REGION Network 2
   RUNG wire#powerrail
      { S7_Templates := "SrcType := Byte" } EQ_Contact(in1 := #Lbyte, in2 := 16#00)
      wire#w1
      Coil( #工作正常 )
   END_RUNG
   RUNG wire#w1
      Coil( #Error.%X1 )
   END_RUNG
   // the same network as SCL:
   #工作正常 := #Lbyte = 16#00;
   #Error.%X1 := #工作正常;
END_REGION

REGION Network 3
   RUNG wire#powerrail
      { S7_Templates := "SrcType := Byte" } EQ_Contact(in1 := #Lbyte, in2 := 16#01)
      wire#w1
      Coil( #无反馈信号 )
   END_RUNG
   RUNG wire#w1
      Coil( #Error.%X2 )
   END_RUNG
   // the same network as SCL:
   #无反馈信号 := #Lbyte = 16#01;
   #Error.%X2 := #无反馈信号;
END_REGION

REGION Network 4
   RUNG wire#powerrail
      { S7_Templates := "SrcType := Byte" } EQ_Contact(in1 := #Lbyte, in2 := 16#02)
      wire#w1
      Coil( #欠压保护 )
   END_RUNG
   RUNG wire#w1
      Coil( #Error.%X3 )
   END_RUNG
   // the same network as SCL:
   #欠压保护 := #Lbyte = 16#02;
   #Error.%X3 := #欠压保护;
END_REGION

REGION Network 5
   RUNG wire#powerrail
      { S7_Templates := "SrcType := Byte" } EQ_Contact(in1 := #Lbyte, in2 := 16#03)
      wire#w1
      Coil( #过压保护 )
   END_RUNG
   RUNG wire#w1
      Coil( #Error.%X4 )
   END_RUNG
   // the same network as SCL:
   #过压保护 := #Lbyte = 16#03;
   #Error.%X4 := #过压保护;
END_REGION

REGION Network 6
   RUNG wire#powerrail
      { S7_Templates := "SrcType := Byte" } EQ_Contact(in1 := #Lbyte, in2 := 16#04)
      wire#w1
      Coil( #过流保护 )
   END_RUNG
   RUNG wire#w1
      Coil( #Error.%X5 )
   END_RUNG
   // the same network as SCL:
   #过流保护 := #Lbyte = 16#04;
   #Error.%X5 := #过流保护;
END_REGION

REGION Network 7
   RUNG wire#powerrail
      { S7_Templates := "SrcType := Byte" } EQ_Contact(in1 := #Lbyte, in2 := 16#05)
      wire#w1
      Coil( #过温保护 )
   END_RUNG
   RUNG wire#w1
      Coil( #Error.%X6 )
   END_RUNG
   // the same network as SCL:
   #过温保护 := #Lbyte = 16#05;
   #Error.%X6 := #过温保护;
END_REGION

REGION Network 8
   RUNG wire#powerrail
      { S7_Templates := "SrcType := Byte" } EQ_Contact(in1 := #Lbyte, in2 := 16#06)
      wire#w1
      Coil( #磁控管故障 )
   END_RUNG
   RUNG wire#w1
      Coil( #Error.%X7 )
   END_RUNG
   // the same network as SCL:
   #磁控管故障 := #Lbyte = 16#06;
   #Error.%X7 := #磁控管故障;
END_REGION

REGION Network 9
   RUNG wire#powerrail
      { S7_Templates := "SrcType := Byte" } EQ_Contact(in1 := #Lbyte, in2 := 16#07)
      wire#w1
      Coil( #浪涌保护 )
   END_RUNG
   RUNG wire#w1
      Coil( #Error.%X8 )
   END_RUNG
   // the same network as SCL:
   #浪涌保护 := #Lbyte = 16#07;
   #Error.%X8 := #浪涌保护;
END_REGION

REGION Network 10
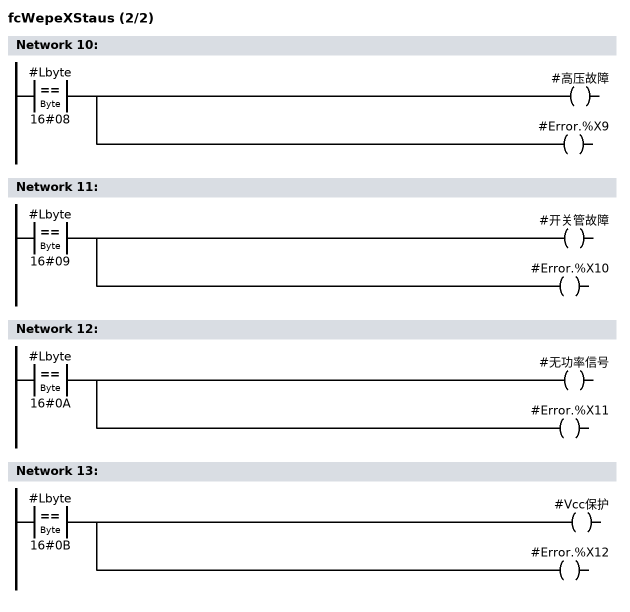
   RUNG wire#powerrail
      { S7_Templates := "SrcType := Byte" } EQ_Contact(in1 := #Lbyte, in2 := 16#08)
      wire#w1
      Coil( #高压故障 )
   END_RUNG
   RUNG wire#w1
      Coil( #Error.%X9 )
   END_RUNG
   // the same network as SCL:
   #高压故障 := #Lbyte = 16#08;
   #Error.%X9 := #高压故障;
END_REGION

REGION Network 11
   RUNG wire#powerrail
      { S7_Templates := "SrcType := Byte" } EQ_Contact(in1 := #Lbyte, in2 := 16#09)
      wire#w1
      Coil( #开关管故障 )
   END_RUNG
   RUNG wire#w1
      Coil( #Error.%X10 )
   END_RUNG
   // the same network as SCL:
   #开关管故障 := #Lbyte = 16#09;
   #Error.%X10 := #开关管故障;
END_REGION

REGION Network 12
   RUNG wire#powerrail
      { S7_Templates := "SrcType := Byte" } EQ_Contact(in1 := #Lbyte, in2 := 16#0A)
      wire#w1
      Coil( #无功率信号 )
   END_RUNG
   RUNG wire#w1
      Coil( #Error.%X11 )
   END_RUNG
   // the same network as SCL:
   #无功率信号 := #Lbyte = 16#0A;
   #Error.%X11 := #无功率信号;
END_REGION

REGION Network 13
   RUNG wire#powerrail
      { S7_Templates := "SrcType := Byte" } EQ_Contact(in1 := #Lbyte, in2 := 16#0B)
      wire#w1
      Coil( #Vcc保护 )
   END_RUNG
   RUNG wire#w1
      Coil( #Error.%X12 )
   END_RUNG
   // the same network as SCL:
   #Vcc保护 := #Lbyte = 16#0B;
   #Error.%X12 := #Vcc保护;
END_REGION
END_FUNCTION

FUNCTION "fcInt_to_mTime" : Void   // FC103, LAD
{ S7_Optimized_Access := 'TRUE' }
VERSION : 0.1
   VAR_INPUT
      intData : Int;
   END_VAR
   VAR_OUTPUT
      mTimeData : Time;
      sTimeData : Time;
   END_VAR
   VAR_TEMP
      dintData1 : DInt;
      dintData2 : DInt;
      dintData3 : DInt;
   END_VAR
BEGIN

REGION Network 1
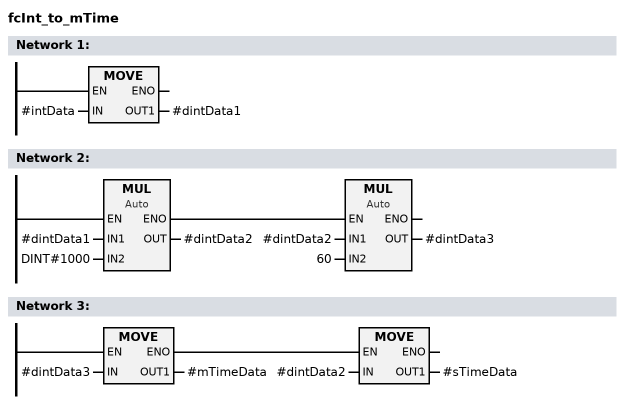
   RUNG wire#powerrail
      Move(in := #intData, out1 => #dintData1)
   END_RUNG
   // the same network as SCL:
   #dintData1 := #intData;
END_REGION

REGION Network 2
   RUNG wire#powerrail
      Mul(in1 := #dintData1, in2 := DINT#1000, out => #dintData2)
      Mul(in1 := #dintData2, in2 := 60, out => #dintData3)
   END_RUNG
   // the same network as SCL:
   #dintData2 := #dintData1 * DINT#1000;
   #dintData3 := #dintData2 * 60;
END_REGION

REGION Network 3
   RUNG wire#powerrail
      Move(in := #dintData3, out1 => #mTimeData)
      Move(in := #dintData2, out1 => #sTimeData)
   END_RUNG
   // the same network as SCL:
   #mTimeData := #dintData3;
   #sTimeData := #dintData2;
END_REGION
END_FUNCTION

FUNCTION "fcArray_Int_mTime" : Void   // FC104, LAD
{ S7_Optimized_Access := 'TRUE' }
VERSION : 0.1
   VAR_INPUT
      "Int" : Array[1..16] of Int;
   END_VAR
   VAR_OUTPUT
      mTimeOut : Array[1..16] of Time;
      sTimeOut : Array[1..16] of Time;
   END_VAR
   VAR_TEMP   // added for the SCL form of the ladder/FBD networks
      _w1 : Bool;
      _w2 : Bool;
      _w3 : Bool;
   END_VAR
BEGIN

REGION Network 1
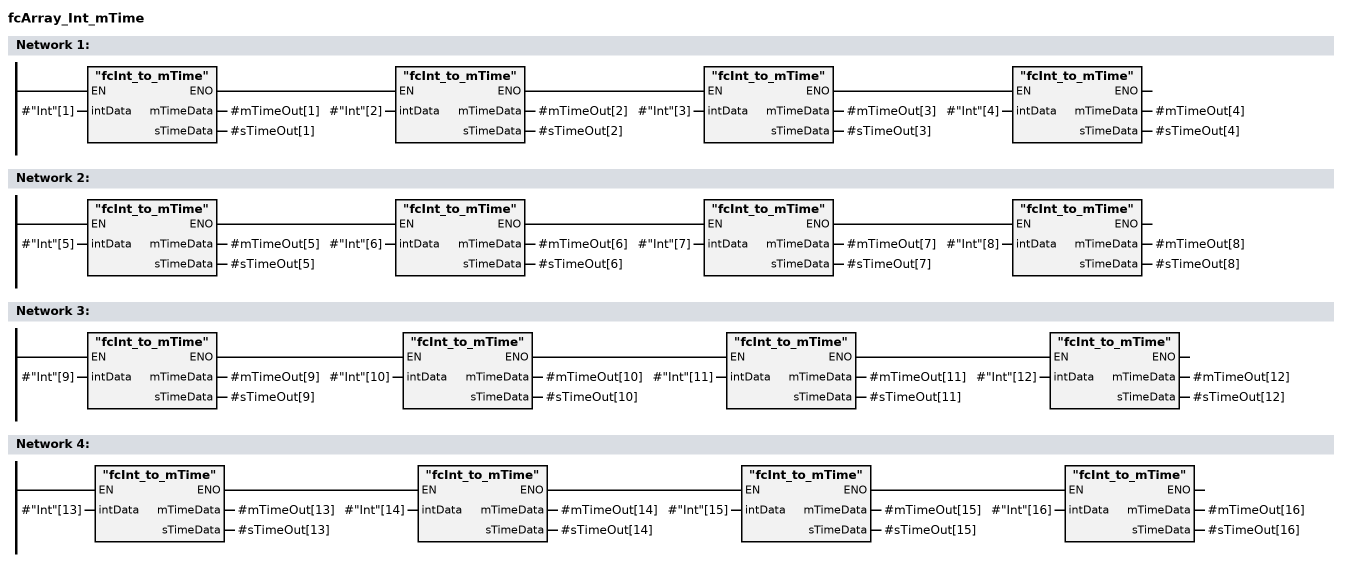
   RUNG wire#powerrail
      "fcInt_to_mTime"(intData := #"Int"[1], mTimeData => #mTimeOut[1], sTimeData => #sTimeOut[1])
      "fcInt_to_mTime"(intData := #"Int"[2], mTimeData => #mTimeOut[2], sTimeData => #sTimeOut[2])
      "fcInt_to_mTime"(intData := #"Int"[3], mTimeData => #mTimeOut[3], sTimeData => #sTimeOut[3])
      "fcInt_to_mTime"(intData := #"Int"[4], mTimeData => #mTimeOut[4], sTimeData => #sTimeOut[4])
   END_RUNG
   // the same network as SCL:
   "fcInt_to_mTime"(intData := #"Int"[1], mTimeData => #mTimeOut[1], sTimeData => #sTimeOut[1], ENO => #_w1);
   "fcInt_to_mTime"(EN := #_w1,
                    intData := #"Int"[2],
                    mTimeData => #mTimeOut[2],
                    sTimeData => #sTimeOut[2],
                    ENO => #_w2);
   "fcInt_to_mTime"(EN := #_w2,
                    intData := #"Int"[3],
                    mTimeData => #mTimeOut[3],
                    sTimeData => #sTimeOut[3],
                    ENO => #_w3);
   IF #_w3 THEN
       "fcInt_to_mTime"(intData := #"Int"[4], mTimeData => #mTimeOut[4], sTimeData => #sTimeOut[4]);
   END_IF;
END_REGION

REGION Network 2
   RUNG wire#powerrail
      "fcInt_to_mTime"(intData := #"Int"[5], mTimeData => #mTimeOut[5], sTimeData => #sTimeOut[5])
      "fcInt_to_mTime"(intData := #"Int"[6], mTimeData => #mTimeOut[6], sTimeData => #sTimeOut[6])
      "fcInt_to_mTime"(intData := #"Int"[7], mTimeData => #mTimeOut[7], sTimeData => #sTimeOut[7])
      "fcInt_to_mTime"(intData := #"Int"[8], mTimeData => #mTimeOut[8], sTimeData => #sTimeOut[8])
   END_RUNG
   // the same network as SCL:
   "fcInt_to_mTime"(intData := #"Int"[5], mTimeData => #mTimeOut[5], sTimeData => #sTimeOut[5], ENO => #_w1);
   "fcInt_to_mTime"(EN := #_w1,
                    intData := #"Int"[6],
                    mTimeData => #mTimeOut[6],
                    sTimeData => #sTimeOut[6],
                    ENO => #_w2);
   "fcInt_to_mTime"(EN := #_w2,
                    intData := #"Int"[7],
                    mTimeData => #mTimeOut[7],
                    sTimeData => #sTimeOut[7],
                    ENO => #_w3);
   IF #_w3 THEN
       "fcInt_to_mTime"(intData := #"Int"[8], mTimeData => #mTimeOut[8], sTimeData => #sTimeOut[8]);
   END_IF;
END_REGION

REGION Network 3
   RUNG wire#powerrail
      "fcInt_to_mTime"(intData := #"Int"[9], mTimeData => #mTimeOut[9], sTimeData => #sTimeOut[9])
      "fcInt_to_mTime"(intData := #"Int"[10], mTimeData => #mTimeOut[10], sTimeData => #sTimeOut[10])
      "fcInt_to_mTime"(intData := #"Int"[11], mTimeData => #mTimeOut[11], sTimeData => #sTimeOut[11])
      "fcInt_to_mTime"(intData := #"Int"[12], mTimeData => #mTimeOut[12], sTimeData => #sTimeOut[12])
   END_RUNG
   // the same network as SCL:
   "fcInt_to_mTime"(intData := #"Int"[9], mTimeData => #mTimeOut[9], sTimeData => #sTimeOut[9], ENO => #_w1);
   "fcInt_to_mTime"(EN := #_w1,
                    intData := #"Int"[10],
                    mTimeData => #mTimeOut[10],
                    sTimeData => #sTimeOut[10],
                    ENO => #_w2);
   "fcInt_to_mTime"(EN := #_w2,
                    intData := #"Int"[11],
                    mTimeData => #mTimeOut[11],
                    sTimeData => #sTimeOut[11],
                    ENO => #_w3);
   IF #_w3 THEN
       "fcInt_to_mTime"(intData := #"Int"[12], mTimeData => #mTimeOut[12], sTimeData => #sTimeOut[12]);
   END_IF;
END_REGION

REGION Network 4
   RUNG wire#powerrail
      "fcInt_to_mTime"(intData := #"Int"[13], mTimeData => #mTimeOut[13], sTimeData => #sTimeOut[13])
      "fcInt_to_mTime"(intData := #"Int"[14], mTimeData => #mTimeOut[14], sTimeData => #sTimeOut[14])
      "fcInt_to_mTime"(intData := #"Int"[15], mTimeData => #mTimeOut[15], sTimeData => #sTimeOut[15])
      "fcInt_to_mTime"(intData := #"Int"[16], mTimeData => #mTimeOut[16], sTimeData => #sTimeOut[16])
   END_RUNG
   // the same network as SCL:
   "fcInt_to_mTime"(intData := #"Int"[13], mTimeData => #mTimeOut[13], sTimeData => #sTimeOut[13], ENO => #_w1);
   "fcInt_to_mTime"(EN := #_w1,
                    intData := #"Int"[14],
                    mTimeData => #mTimeOut[14],
                    sTimeData => #sTimeOut[14],
                    ENO => #_w2);
   "fcInt_to_mTime"(EN := #_w2,
                    intData := #"Int"[15],
                    mTimeData => #mTimeOut[15],
                    sTimeData => #sTimeOut[15],
                    ENO => #_w3);
   IF #_w3 THEN
       "fcInt_to_mTime"(intData := #"Int"[16], mTimeData => #mTimeOut[16], sTimeData => #sTimeOut[16]);
   END_IF;
END_REGION
END_FUNCTION

FUNCTION "fcArray_bool_to_bool" : Void   // FC105, LAD
{ S7_Optimized_Access := 'TRUE' }
VERSION : 0.1
   VAR_INPUT
      In : Array[1..16] of Bool;
   END_VAR
   VAR_OUTPUT
      Out : Bool;
   END_VAR
BEGIN

REGION Network 1
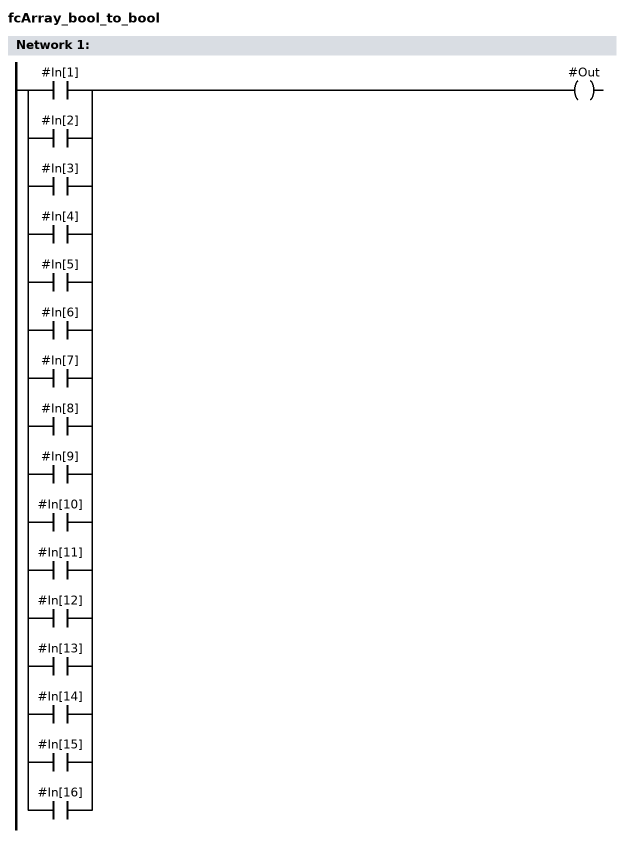
   RUNG wire#powerrail
      Contact( #In[1] )
      wire#w1
      Coil( #Out )
   END_RUNG
   RUNG wire#powerrail
      Contact( #In[2] )
   END_RUNG wire#w1
   RUNG wire#powerrail
      Contact( #In[3] )
   END_RUNG wire#w1
   RUNG wire#powerrail
      Contact( #In[4] )
   END_RUNG wire#w1
   RUNG wire#powerrail
      Contact( #In[5] )
   END_RUNG wire#w1
   RUNG wire#powerrail
      Contact( #In[6] )
   END_RUNG wire#w1
   RUNG wire#powerrail
      Contact( #In[7] )
   END_RUNG wire#w1
   RUNG wire#powerrail
      Contact( #In[8] )
   END_RUNG wire#w1
   RUNG wire#powerrail
      Contact( #In[9] )
   END_RUNG wire#w1
   RUNG wire#powerrail
      Contact( #In[10] )
   END_RUNG wire#w1
   RUNG wire#powerrail
      Contact( #In[11] )
   END_RUNG wire#w1
   RUNG wire#powerrail
      Contact( #In[12] )
   END_RUNG wire#w1
   RUNG wire#powerrail
      Contact( #In[13] )
   END_RUNG wire#w1
   RUNG wire#powerrail
      Contact( #In[14] )
   END_RUNG wire#w1
   RUNG wire#powerrail
      Contact( #In[15] )
   END_RUNG wire#w1
   RUNG wire#powerrail
      Contact( #In[16] )
   END_RUNG wire#w1
   // the same network as SCL:
   #Out := #In[1] OR #In[2] OR #In[3] OR #In[4] OR #In[5] OR #In[6] OR #In[7] OR #In[8] OR #In[9] OR #In[10] OR #In[11] OR #In[12] OR #In[13] OR #In[14] OR #In[15] OR #In[16];
END_REGION
END_FUNCTION

ORGANIZATION_BLOCK "Main"   // OB1, LAD, ProgramCycle
TITLE = "Main Program Sweep (Cycle)"
{ S7_Optimized_Access := 'TRUE' }
VERSION : 0.1
   VAR_INPUT
      Initial_Call : Bool;   // Initial call of this OB
      Remanence : Bool;   // =True, if remanent data are available
   END_VAR
BEGIN

REGION Network 1
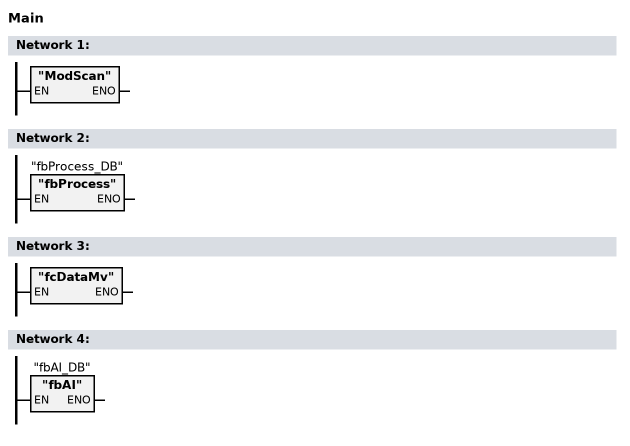
   RUNG wire#powerrail
      "ModScan"()
   END_RUNG
   // the same network as SCL:
   "ModScan"();
END_REGION

REGION Network 2
   RUNG wire#powerrail
      "fbProcess_DB"()
   END_RUNG
   // the same network as SCL:
   "fbProcess_DB"();   // "fbProcess"
END_REGION

REGION Network 3
   RUNG wire#powerrail
      "fcDataMv"()
   END_RUNG
   // the same network as SCL:
   "fcDataMv"();
END_REGION

REGION Network 4
   RUNG wire#powerrail
      "fbAI_DB"()
   END_RUNG
   // the same network as SCL:
   "fbAI_DB"();   // "fbAI"
END_REGION
END_ORGANIZATION_BLOCK

// folder: System blocks/Program resources

FUNCTION "ModScan" : Void   // FC10000, LAD
TITLE = ModScan
{ S7_Optimized_Access := 'TRUE' }
AUTHOR : SIMATIC
VERSION : 4.0
BEGIN

REGION Network 1: Modbus-RTU Job scan
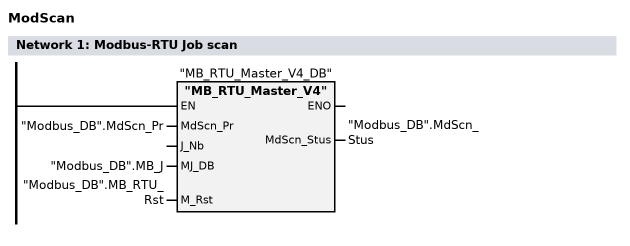
   RUNG wire#powerrail
      "MB_RTU_Master_V4_DB"(MdScn_Pr := "Modbus_DB".MdScn_Pr, J_Nb :=, MJ_DB := "Modbus_DB".MB_J, M_Rst := "Modbus_DB".MB_RTU_Rst, MdScn_Stus => "Modbus_DB".MdScn_Stus)
   END_RUNG
   // the same network as SCL:
   "MB_RTU_Master_V4_DB"(MdScn_Pr := "Modbus_DB".MdScn_Pr,   // "MB_RTU_Master_V4"
                         MJ_DB := "Modbus_DB".MB_J,
                         M_Rst := "Modbus_DB".MB_RTU_Rst,
                         MdScn_Stus => "Modbus_DB".MdScn_Stus);
END_REGION
END_FUNCTION

(* ===== HMI "HMI_RT_1" =====
system functions are stored by id; their names below are inferred from use
connection "HMI_连接_1": ETHERNET, SMART_S7_1200_OMS

HMI tags "变量表_1"
   "WepeX_PowerSPCom" : Int = PLC dbHMI.WepeX_PowerSPCom AT %DB50.DBW0, 1 s
   "WepeX_ActpowerCom" : Int = PLC dbHMI.WepeX_ActpowerCom AT %DB50.DBW38, 1 s
   "Mode" : Bool = PLC dbHMI.Mode AT %DB50.DBX164.0, 1 s
   "WepeX_PowerMan" : Bool = PLC dbHMI.WepeX_PowerMan AT %DB50.DBX164.1, 1 s
   "CoolingWaterMan" : Bool = PLC dbHMI.CoolingWaterMan AT %DB50.DBX164.2, 1 s
   "AirCompressorMan" : Bool = PLC dbHMI.AirCompressorMan AT %DB50.DBX164.3, 1 s
   "BlowerMan" : Bool = PLC dbHMI.BlowerMan AT %DB50.DBX164.4, 1 s
   "PeristalticpumpMan" : Bool = PLC dbHMI.PeristalticpumpMan AT %DB50.DBX164.5, 1 s
   "1YV1Man" : Bool = PLC dbHMI.1YV1Man AT %DB50.DBX164.6, 1 s
   "1YV2Man" : Bool = PLC dbHMI.1YV2Man AT %DB50.DBX164.7, 1 s
   "2YV1Man" : Bool = PLC dbHMI.2YV1Man AT %DB50.DBX165.0, 1 s
   "2YV2Man" : Bool = PLC dbHMI.2YV2Man AT %DB50.DBX165.1, 1 s
   "WepeXP1通信正常" : Bool = PLC dbHMI.WepeXP1通信正常 AT %DB50.DBX170.0, 1 s
   "WepeXP1通信不正常" : Bool = PLC dbHMI.WepeXP1通信不正常 AT %DB50.DBX170.1, 1 s
   "WepeXP1工作正常" : Bool = PLC dbHMI.WepeXP1工作正常 AT %DB50.DBX170.2, 1 s
   "WepeXP1无反馈信号" : Bool = PLC dbHMI.WepeXP1无反馈信号 AT %DB50.DBX170.3, 1 s
   "WepeXP1欠压保护" : Bool = PLC dbHMI.WepeXP1欠压保护 AT %DB50.DBX170.4, 1 s
   "WepeXP1过压保护" : Bool = PLC dbHMI.WepeXP1过压保护 AT %DB50.DBX170.5, 1 s
   "WepeXP1过流保护" : Bool = PLC dbHMI.WepeXP1过流保护 AT %DB50.DBX170.6, 1 s
   "WepeXP1过温保护" : Bool = PLC dbHMI.WepeXP1过温保护 AT %DB50.DBX170.7, 1 s
   "WepeXP1磁控管故障" : Bool = PLC dbHMI.WepeXP1磁控管故障 AT %DB50.DBX171.0, 1 s
   "WepeXP1浪涌保护" : Bool = PLC dbHMI.WepeXP1浪涌保护 AT %DB50.DBX171.1, 1 s
   "WepeXP1高压故障" : Bool = PLC dbHMI.WepeXP1高压故障 AT %DB50.DBX171.2, 1 s
   "WepeXP1开关管故障" : Bool = PLC dbHMI.WepeXP1开关管故障 AT %DB50.DBX171.3, 1 s
   "WepeXP1无功率信号" : Bool = PLC dbHMI.WepeXP1无功率信号 AT %DB50.DBX171.4, 1 s
   "WepeXP1Vcc保护" : Bool = PLC dbHMI.WepeXP1Vcc保护 AT %DB50.DBX171.5, 1 s
   "WepeXP1通信状态" : Int = PLC dbHMI.WepeXP1通信状态 AT %DB50.DBW172, 1 s
   "微波状态" : Int = PLC dbHMI.微波状态 AT %DB50.DBW174, 1 s
   "火炬状态" : Int = PLC dbHMI.火炬状态 AT %DB50.DBW176, 1 s
   "Start" : Bool = PLC dbHMI.Start AT %DB50.DBX178.0, 1 s
   "Stop" : Bool = PLC dbHMI.Stop AT %DB50.DBX178.1, 1 s
   "Reset" : Bool = PLC dbHMI.Reset AT %DB50.DBX178.2, 1 s
   "Running" : Bool = PLC dbHMI.Running AT %DB50.DBX178.3, 1 s
   "WepeXPowerOut" : Bool = PLC WepeXEnable AT %Q0.1, 1 s
   "CoolingWater" : Bool = PLC CoolingWater AT %Q0.2, 1 s
   "Blower" : Bool = PLC Blower AT %Q0.3, 1 s
   "AirCompressor" : Bool = PLC AirCompressor AT %Q0.4, 1 s
   "Peristalticpump" : Bool = PLC Peristalticpump AT %Q0.0, 1 s
   "气体温度" : Real = PLC dbHMI.气体温度 AT %DB50.DBD180, 1 s
   "1YV1" : Bool = PLC 1YV1 AT %Q1.0, 1 s
   "1YV2" : Bool = PLC 1YV2 AT %Q1.1, 1 s
   "2YV1" : Bool = PLC 2YV1 AT %Q1.2, 1 s
   "2YV2" : Bool = PLC 2YV2 AT %Q1.3, 1 s
   "3YV1Man" : Bool = PLC dbHMI.3YV1Man AT %DB50.DBX165.2, 1 s
   "3YV1" : Bool = PLC 3YV1 AT %Q1.4, 1 s
   "3YV2Man" : Bool = PLC dbHMI.3YV2Man AT %DB50.DBX165.3, 1 s
   "3YV2" : Bool = PLC 3YV2 AT %Q1.5, 1 s
   "4YVMan" : Bool = PLC dbHMI.4YVMan AT %DB50.DBX165.4, 1 s
   "4YV" : Bool = PLC 4YV AT %Q1.6, 1 s
   "inUnit.Coolingwater" : Bool = PLC dbHMI.inUnit.Coolingwater AT %DB50.DBX184.0, 1 s
   "inUnit.AirCompressor" : Bool = PLC dbHMI.inUnit.AirCompressor AT %DB50.DBX184.1, 1 s
   "inUnit.Peristalticpump" : Bool = PLC dbHMI.inUnit.Peristalticpump AT %DB50.DBX184.2, 1 s
   "inUnit.WepeX_Enable" : Bool = PLC dbHMI.inUnit.WepeX_Enable AT %DB50.DBX184.3, 1 s
   "inUnit.AYV1" : Bool = PLC dbHMI.inUnit.AYV1 AT %DB50.DBX184.4, 1 s
   "inUnit.AYV2" : Bool = PLC dbHMI.inUnit.AYV2 AT %DB50.DBX184.5, 1 s
   "inUnit.BYV1" : Bool = PLC dbHMI.inUnit.BYV1 AT %DB50.DBX184.6, 1 s
   "inUnit.BYV2" : Bool = PLC dbHMI.inUnit.BYV2 AT %DB50.DBX184.7, 1 s
   "inUnit.CYV1" : Bool = PLC dbHMI.inUnit.CYV1 AT %DB50.DBX185.0, 1 s
   "inUnit.CYV2" : Bool = PLC dbHMI.inUnit.CYV2 AT %DB50.DBX185.1, 1 s
   "inUnit.DYV" : Bool = PLC dbHMI.inUnit.DYV AT %DB50.DBX185.2, 1 s
   "inUnit.Blower" : Bool = PLC dbHMI.inUnit.Blower AT %DB50.DBX185.3, 1 s
   "inUnit.Runtime" : Int = PLC dbHMI.inUnit.Runtime AT %DB50.DBW186, 1 s
   "inUnit.WepeX_Power" : Int = PLC dbHMI.inUnit.WepeX_Power AT %DB50.DBW188, 1 s
   "inUnit.Donebit" : Int = PLC dbHMI.inUnit.Donebit AT %DB50.DBW190, 1 s
   "ActUnit.Coolingwater" : Bool = PLC dbHMI.ActRcpUnit.Coolingwater AT %DB50.DBX202.0, 1 s
   "ActUnit.AirCompressor" : Bool = PLC dbHMI.ActRcpUnit.AirCompressor AT %DB50.DBX202.1, 1 s
   "ActUnit.Peristalticpump" : Bool = PLC dbHMI.ActRcpUnit.Peristalticpump AT %DB50.DBX202.2, 1 s
   "ActUnit.WepeX_Enable" : Bool = PLC dbHMI.ActRcpUnit.WepeX_Enable AT %DB50.DBX202.3, 1 s
   "ActUnit.AYV1" : Bool = PLC dbHMI.ActRcpUnit.AYV1 AT %DB50.DBX202.4, 1 s
   "ActUnit.AYV2" : Bool = PLC dbHMI.ActRcpUnit.AYV2 AT %DB50.DBX202.5, 1 s
   "ActUnit.BYV1" : Bool = PLC dbHMI.ActRcpUnit.BYV1 AT %DB50.DBX202.6, 1 s
   "ActUnit.BYV2" : Bool = PLC dbHMI.ActRcpUnit.BYV2 AT %DB50.DBX202.7, 1 s
   "ActUnit.CYV1" : Bool = PLC dbHMI.ActRcpUnit.CYV1 AT %DB50.DBX203.0, 1 s
   "ActUnit.CYV2" : Bool = PLC dbHMI.ActRcpUnit.CYV2 AT %DB50.DBX203.1, 1 s
   "ActUnit.DYV" : Bool = PLC dbHMI.ActRcpUnit.DYV AT %DB50.DBX203.2, 1 s
   "ActUnit.Blower" : Bool = PLC dbHMI.ActRcpUnit.Blower AT %DB50.DBX203.3, 1 s
   "ActUnit.Runtime" : Int = PLC dbHMI.ActRcpUnit.Runtime AT %DB50.DBW204, 1 s
   "ActUnit.WepeX_Power" : Int = PLC dbHMI.ActRcpUnit.WepeX_Power AT %DB50.DBW206, 1 s
   "ActUnit.Donebit" : Int = PLC dbHMI.ActRcpUnit.Donebit AT %DB50.DBW208, 1 s
   "RecipeNum" : Int = PLC dbHMI.RecipeNum AT %DB50.DBW192, 1 s
   "StepNumMan" : Int = PLC dbHMI.StepNumMan AT %DB50.DBW194, 1 s
   "Editor" : Bool = PLC dbHMI.Editor AT %DB50.DBX200.0, 1 s
   "Save" : Bool = PLC dbHMI.Save AT %DB50.DBX200.1, 1 s

discrete alarms
   1: '', class Errors

Template "模板_1" 800x480
   Button "模板_按钮_1" at 0,448 size 96x32; TextOff '自动页面'
      on Click: ActivateScreen("1自动画面", 0)
   Button "模板_按钮_2" at 96,448 size 96x32; TextOff '手动页面'
      on Click: ActivateScreen("2手动画面", 0)
   Button "模板_按钮_3" at 192,448 size 96x32; TextOff '程序设置'
      on Click: ActivateScreen("3程序设置", 0)
   Button "模板_按钮_4" at 288,448 size 96x32; TextOff '温度曲线'
      on Click: ActivateScreen("4温度曲线", 0)
   Button "模板_按钮_5" at 384,448 size 96x32; TextOff '报警信息'
      Appearance <- "Mode"
      on Click: ActivateScreen("5报警信息", 0)
   Button "模板_按钮_6" at 480,448 size 96x32; TextOff '自/手模式'
      on Press: InvertBit("Mode")
      Appearance <- "Mode"

screen "1自动画面" 800x480, template "模板_1"
   TextField "文本域_16" at 73,86 size 57x16; Text '设备状态'
   TextField "文本域_17" at 103,145 size 31x16; Text '微波'
   TextField "文本域_18" at 103,177 size 31x16; Text '火炬'
   TextField "文本域_19" at 103,113 size 31x16; Text '通信'
   TextField "文本域_20" at 102,211 size 31x16; Text '过流'
   TextField "文本域_21" at 102,245 size 31x16; Text '欠流'
   TextField "文本域_22" at 102,280 size 31x16; Text '超温'
   TextField "文本域_14" at 325,75 size 73x20; Text '程序选择'
   Button "按钮_1" at 316,114 size 97x32; TextOff '开放式'
   Button "按钮_2" at 316,187 size 97x32; TextOff '管道式'
   Button "按钮_3" at 314,259 size 97x32; TextOff '自定义'
   Button "按钮_7" at 153,343 size 81x70; TextOff '启动'
      on Press: SetBit("Start")
      on Release: ResetBit("Start")
      Appearance <- "Running"
   TextField "文本域_6" at 575,199 size 73x20; Text '气体余量'
   IOField "I/O 域_4" at 646,191 size 96x32; FormatPattern 9999999
   TextField "文本域_7" at 576,95 size 73x20; Text '实际功率'
   IOField "I/O 域_5" at 648,90 size 96x32; FormatPattern s99999
      ProcessValue <- "WepeX_ActpowerCom"
   TextField "文本域_8" at 745,94 size 16x23; Text 'W'
   TextField "文本域_9" at 575,149 size 73x20; Text '气体温度'
   IOField "I/O 域_6" at 648,141 size 96x32; FormatPattern s999.99
      ProcessValue <- "气体温度"
   TextField "文本域_10" at 745,147 size 25x23; Text '℃'
   Button "按钮_8" at 382,348 size 80x68; TextOff '停止'
      on Press: SetBit("Stop")
      on Release: ResetBit("Stop")
   TextField "文本域_1" at 237,14 size 275x33; Text '多功能等离子消毒机'
   Circle "圆_1" at 74,112 size 20x20
      Appearance <- "WepeXP1通信不正常"
   Circle "圆_2" at 74,144 size 20x20
      Appearance <- "微波状态"
   Circle "圆_3" at 74,177 size 20x20
      Appearance <- "火炬状态"
   Circle "圆_4" at 74,210 size 20x20
      Appearance <- "WepeXP1过流保护"
   Circle "圆_5" at 74,243 size 20x20
      Appearance <- "WepeXP1欠压保护"
   Circle "圆_6" at 74,277 size 20x20
      Appearance <- "WepeXP1过温保护"
   Button "按钮_9" at 606,349 size 82x64; TextOff '复位'
      on Press: SetBit("Reset")
      on Release: ResetBit("Reset")
   TextField "文本域_4" at 749,197 size 16x23; Text '%'

screen "2手动画面" 800x480, template "模板_1"
   Button "按钮_1" at 169,84 size 80x55; TextOff '冷水机'
      on Press: InvertBit("CoolingWaterMan")
      Appearance <- "CoolingWaterMan"
   Button "按钮_2" at 169,258 size 80x55; TextOff '空压机'
      on Press: InvertBit("AirCompressorMan")
      Appearance <- "AirCompressorMan"
   Button "按钮_3" at 169,170 size 80x55; TextOff '风机'
      on Press: InvertBit("BlowerMan")
      Appearance <- "BlowerMan"
   Button "按钮_4" at 169,348 size 80x55; TextOff '蠕动泵'
      on Press: InvertBit("PeristalticpumpMan")
      Appearance <- "PeristalticpumpMan"
   TextField "文本域_6" at 617,102 size 73x20; Text '功率设置'
   IOField "I/O 域_4" at 697,95 size 64x32; FormatPattern 9999
      ProcessValue <- "WepeX_PowerSPCom"
   TextField "文本域_7" at 620,156 size 73x20; Text '实际功率'
   IOField "I/O 域_5" at 700,149 size 57x32; FormatPattern 9999
      ProcessValue <- "WepeX_ActpowerCom"
   TextField "文本域_8" at 764,154 size 16x23; Text 'W'
   TextField "文本域_9" at 620,210 size 73x20; Text '气体余量'
   IOField "I/O 域_6" at 695,205 size 63x32; FormatPattern 999
   TextField "文本域_10" at 755,269 size 25x23; Text '℃'
   TextField "文本域_1" at 763,98 size 16x23; Text 'W'
   Button "按钮_5" at 333,82 size 80x55; TextOff '功率'
      on Press: InvertBit("WepeX_PowerMan")
      Appearance <- "WepeX_PowerMan"
   Button "按钮_6" at 490,83 size 80x55; TextOff '阀门进1'
      on Press: InvertBit("1YV1Man")
      Appearance <- "1YV1Man"
   Button "按钮_7" at 490,170 size 80x55; TextOff '阀门进2'
      on Press: InvertBit("1YV2Man")
      Appearance <- "1YV2Man"
   Button "按钮_8" at 488,259 size 80x55; TextOff '阀门出1'
      on Press: InvertBit("2YV1Man")
      Appearance <- "2YV1Man"
   Button "按钮_9" at 490,345 size 80x55; TextOff '阀门出2'
      on Press: InvertBit("2YV2Man")
      Appearance <- "2YV2Man"
   Circle "圆_8" at 258,100 size 20x20
      Appearance <- "CoolingWater"
   Circle "圆_9" at 256,275 size 20x20
      Appearance <- "AirCompressor"
   Circle "圆_10" at 257,189 size 20x20
      Appearance <- "Blower"
   Circle "圆_11" at 257,362 size 20x20
      Appearance <- "Peristalticpump"
   Circle "圆_12" at 417,100 size 20x20
      Appearance <- "WepeXPowerOut"
   Circle "圆_13" at 575,103 size 20x20
      Appearance <- "1YV1"
   Circle "圆_14" at 573,188 size 20x20
      Appearance <- "1YV2"
   Circle "圆_15" at 570,275 size 20x20
      Appearance <- "2YV1"
   Circle "圆_16" at 573,363 size 20x20
      Appearance <- "2YV2"
   Button "按钮_10" at 333,258 size 80x55; TextOff '氮气阀1'
      on Press: InvertBit("3YV1Man")
      Appearance <- "3YV1Man"
   Circle "圆_17" at 416,272 size 20x20
      Appearance <- "3YV1"
   Button "按钮_11" at 333,344 size 80x55; TextOff '氮气阀2'
      on Press: InvertBit("3YV2Man")
      Appearance <- "3YV2Man"
   Circle "圆_18" at 416,359 size 20x20
      Appearance <- "3YV2"
   Button "按钮_12" at 333,170 size 80x55; TextOff '氧气阀'
      on Press: InvertBit("4YVMan")
      Appearance <- "4YVMan"
   Circle "圆_19" at 417,186 size 20x20
      Appearance <- "4YV"
   TextField "文本域_16" at 43,120 size 57x16; Text '设备状态'
   TextField "文本域_17" at 73,179 size 31x16; Text '微波'
   TextField "文本域_18" at 73,211 size 31x16; Text '火炬'
   TextField "文本域_19" at 73,147 size 31x16; Text '通信'
   TextField "文本域_20" at 72,245 size 31x16; Text '过流'
   TextField "文本域_21" at 72,279 size 31x16; Text '欠流'
   TextField "文本域_22" at 72,314 size 31x16; Text '超温'
   Circle "圆_1" at 44,146 size 20x20
      Appearance <- "WepeXP1通信不正常"
   Circle "圆_2" at 44,178 size 20x20
      Appearance <- "微波状态"
   Circle "圆_3" at 44,211 size 20x20
      Appearance <- "火炬状态"
   Circle "圆_4" at 44,244 size 20x20
      Appearance <- "WepeXP1过流保护"
   Circle "圆_5" at 44,277 size 20x20
      Appearance <- "WepeXP1欠压保护"
   Circle "圆_6" at 44,311 size 20x20
      Appearance <- "WepeXP1过温保护"
   TextField "文本域_2" at 763,208 size 16x23; Text '%'
   TextField "文本域_3" at 618,269 size 73x20; Text '气体温度'
   IOField "I/O 域_1" at 694,264 size 58x32; FormatPattern 999
      ProcessValue <- "气体温度"
   TextField "文本域_4" at 237,14 size 275x33; Text '多功能等离子消毒机'

screen "3程序设置" 800x480, template "模板_1"
   TextField "文本域_2" at 330,28 size 109x29; Text '程序编辑'
   Button "按钮_1" at 250,126 size 80x40; TextOff '冷水机'
      on Press: InvertBit("inUnit.Coolingwater")
      Appearance <- "inUnit.Coolingwater"
   Button "按钮_2" at 430,128 size 80x40; TextOff '空压机'
      on Press: InvertBit("inUnit.AirCompressor")
      Appearance <- "inUnit.AirCompressor"
   Button "按钮_3" at 250,187 size 80x40; TextOff '风机'
      on Press: InvertBit("inUnit.Blower")
      Appearance <- "inUnit.Blower"
   Button "按钮_4" at 430,186 size 80x40; TextOff '蠕动泵'
      on Press: InvertBit("inUnit.Peristalticpump")
      Appearance <- "inUnit.Peristalticpump"
   Button "按钮_5" at 428,247 size 80x40; TextOff '功率'
      on Press: InvertBit("ActUnit.WepeX_Enable")
      Appearance <- "inUnit.WepeX_Enable"
   Button "按钮_6" at 606,186 size 80x40; TextOff '阀门进1'
      on Press: InvertBit("inUnit.AYV1")
      Appearance <- "inUnit.AYV1"
   Button "按钮_7" at 607,249 size 80x40; TextOff '阀门进2'
      on Press: InvertBit("inUnit.AYV2")
      Appearance <- "inUnit.AYV2"
   Button "按钮_8" at 606,307 size 80x40; TextOff '阀门出1'
      on Press: InvertBit("inUnit.BYV1")
      Appearance <- "inUnit.BYV1"
   Button "按钮_9" at 606,368 size 80x40; TextOff '阀门出2'
      on Press: InvertBit("inUnit.BYV2")
      Appearance <- "inUnit.BYV2"
   Circle "圆_8" at 358,131 size 32x32
      Appearance <- "ActUnit.Coolingwater"
   Circle "圆_9" at 538,130 size 32x32
      Appearance <- "ActUnit.AirCompressor"
   Circle "圆_10" at 358,191 size 32x32
      Appearance <- "ActUnit.Blower"
   Circle "圆_11" at 537,190 size 32x32
      Appearance <- "ActUnit.Peristalticpump"
   Circle "圆_12" at 541,251 size 32x32
      Appearance <- "ActUnit.WepeX_Enable"
   Circle "圆_13" at 719,188 size 32x32
      Appearance <- "ActUnit.AYV1"
   Circle "圆_14" at 719,253 size 32x32
      Appearance <- "ActUnit.AYV2"
   Circle "圆_15" at 718,310 size 32x32
      Appearance <- "ActUnit.BYV1"
   Circle "圆_16" at 719,368 size 32x32
      Appearance <- "ActUnit.BYV2"
   Button "按钮_10" at 427,309 size 80x40; TextOff '氮气阀1'
      on Press: InvertBit("inUnit.CYV1")
      Appearance <- "inUnit.CYV1"
   Circle "圆_17" at 540,312 size 32x32
      Appearance <- "ActUnit.CYV1"
   Button "按钮_11" at 427,369 size 80x40; TextOff '氮气阀2'
      on Press: InvertBit("inUnit.CYV2")
      Appearance <- "inUnit.CYV2"
   Circle "圆_18" at 542,371 size 32x32
      Appearance <- "ActUnit.CYV2"
   Button "按钮_12" at 607,127 size 80x40; TextOff '氧气阀'
      on Press: InvertBit("inUnit.DYV")
      Appearance <- "inUnit.DYV"
   Circle "圆_19" at 718,131 size 32x32
      Appearance <- "ActUnit.DYV"
   TextField "文本域_6" at 40,72 size 71x25; Text '程序号'
   IOField "I/O 域_4" at 143,69 size 64x32; FormatPattern 9999
      ProcessValue <- "RecipeNum"
   TextField "文本域_1" at 38,121 size 71x25; Text '步序号'
   IOField "I/O 域_1" at 142,115 size 64x32; FormatPattern 9999
      ProcessValue <- "StepNumMan"
   Button "按钮_13" at 77,320 size 80x40; TextOff '编辑'
      on Press: InvertBit("Editor")
      Appearance <- "AirCompressorMan"
   Button "按钮_14" at 79,378 size 80x40; TextOff '保存'
      on Press: SetBit("Save")
      Appearance <- "AirCompressorMan"
      on Release: ResetBit("Save")
   TextField "文本域_3" at 248,77 size 93x25; Text '设备单元'
   TextField "文本域_4" at 422,78 size 93x25; Text '设备单元'
   TextField "文本域_5" at 602,79 size 93x25; Text '设备单元'
   TextField "文本域_7" at 355,79 size 49x25; Text '状态'
   TextField "文本域_8" at 530,79 size 49x25; Text '状态'
   TextField "文本域_9" at 711,79 size 49x25; Text '状态'
   TextField "文本域_10" at 34,171 size 93x25; Text '步序时间'
   IOField "I/O 域_2" at 140,165 size 72x32; FormatPattern 99999
      ProcessValue <- "inUnit.Runtime"
   TextField "文本域_11" at 40,273 size 93x25; Text '结束标识'
   IOField "I/O 域_3" at 141,269 size 64x32; FormatPattern 9
      ProcessValue <- "inUnit.Donebit"
   TextField "文本域_13" at 249,364 size 42x25; Text '结束'
   IOField "I/O 域_6" at 315,374 size 64x32; FormatPattern 9999
      ProcessValue <- "ActUnit.Donebit"
   TextField "文本域_14" at 249,387 size 41x21; Text '标识'
   TextField "文本域_15" at 250,304 size 42x25; Text '当前'
   TextField "文本域_16" at 251,327 size 41x21; Text '时间'
   TextField "文本域_17" at 251,244 size 42x25; Text '微波'
   TextField "文本域_18" at 251,267 size 41x21; Text '功率'
   IOField "I/O 域_7" at 314,312 size 71x32; FormatPattern 99999
      ProcessValue <- "ActUnit.Runtime"
   IOField "I/O 域_8" at 315,251 size 64x32; FormatPattern 9999
      ProcessValue <- "WepeX_PowerSPCom"
   TextField "文本域_12" at 382,256 size 16x23; Text 'W'
   TextField "文本域_19" at 386,316 size 16x23; Text 'S'
   TextField "文本域_20" at 35,221 size 93x25; Text '微波功率'
   IOField "I/O 域_5" at 143,214 size 64x32; FormatPattern 9999
      ProcessValue <- "inUnit.WepeX_Power"
   TextField "文本域_21" at 209,220 size 16x23; Text 'W'
   TextField "文本域_22" at 212,170 size 16x23; Text 'S'

screen "4温度曲线" 800x480, template "模板_1"
   TrendView "趋势视图_1" at 91,67 size 600x300

screen "5报警信息" 800x480, template "模板_1"
   AlarmView "报警视图_1" at 89,64 size 593x324
*)